
   //******************************************************************************************************
   #q_byDriveState := WORD_TO_BYTE(#ILx2T_Ref.i_woDriveStatus AND 16#000F);
   #q_xReadyToSwitchOn := #q_byDriveState = 4;
   #q_xSwitchedOn := #q_byDriveState = 6 OR #q_byDriveState = 7;
   #q_xFault := #ILx2T_Ref.stDriveStatus.FaultActive;
   #q_xWarning := #ILx2T_Ref.stDriveStatus.WarningActive;
   #q_xHALT_active := #ILx2T_Ref.stDriveStatus.HaltActive;
   #q_xRef_OK := #ILx2T_Ref.i_by_ModeStatus.%X5;
   #q_xQuickStop_Active := (#q_byDriveState = 7) AND #ILx2T_Ref.stDriveStatus.x_End;
   //******************************************************************************************************
   // MotionStat
   #q_xStandstill := #ILx2T_Ref.stDriveStatus.x_End;
   #q_xPositiveDirection := #ILx2T_Ref.i_wo_ActionWord.%X7;
   #q_xNegativeDirection := #ILx2T_Ref.i_wo_ActionWord.%X8;
   //#q_xInPositionWindow := #ILx2T_Ref.i_wo_ActionWord.%X9;
   #q_xTargetVelocityZero := #ILx2T_Ref.i_wo_ActionWord.%X11;
   #q_xAccelerating := #ILx2T_Ref.i_wo_ActionWord.%X13;
   #q_xDecelerating := #ILx2T_Ref.i_wo_ActionWord.%X12;
   #q_xConstantVelocity := #ILx2T_Ref.i_wo_ActionWord.%X14;

   #ILx2T_Ref.st_ActionWord.MotionNegative := #q_xNegativeDirection;
   //#ILx2T_Ref.st_ActionWord.InsidePosWindow := #q_xInPositionWindow;
   #ILx2T_Ref.st_ActionWord.TargetVelocityZero := #q_xTargetVelocityZero;
   #ILx2T_Ref.st_ActionWord.Decelerating := #q_xDecelerating;
   #ILx2T_Ref.st_ActionWord.Accelerating := #q_xAccelerating;
   #ILx2T_Ref.st_ActionWord.ConstantVelocity := #q_xConstantVelocity;
   #ILx2T_Ref.st_ActionWord.MotionZero := #q_xStandstill;
   #ILx2T_Ref.st_ActionWord.MotionPositive := #q_xPositiveDirection;;

   //******************************************************************************************************
   // digital Drive Inputs
   #ILx2T_Ref.x_IO_1 := #ILx2T_Ref.i_by_driveInput.%X0;
   #ILx2T_Ref.x_IO_2 := #ILx2T_Ref.i_by_driveInput.%X1;
   #ILx2T_Ref.x_IO_3 := #ILx2T_Ref.i_by_driveInput.%X2;
   #ILx2T_Ref.x_IO_4 := #ILx2T_Ref.i_by_driveInput.%X3;
   #ILx2T_Ref.x_STO_A := #ILx2T_Ref.i_by_driveInput.%X4;
   #ILx2T_Ref.x_STO_B := #ILx2T_Ref.i_by_driveInput.%X5;
   //******************************************************************************************************
   // mfStat
   #ILx2T_Ref.by_OP_ModeAct := #ILx2T_Ref.i_by_ModeStatus AND 16#0F;

   #ILx2T_Ref.st_ModeStatus.Reference_OK := #ILx2T_Ref.i_by_ModeStatus.%X5;
   #q_xRef_OK := #ILx2T_Ref.st_ModeStatus.Reference_OK;
   #ILx2T_Ref.st_ModeStatus.ModeError := #ILx2T_Ref.i_by_ModeStatus.%X6;
   #ILx2T_Ref.st_ModeStatus.ModeToggle := #ILx2T_Ref.i_by_ModeStatus.%X7;

   //******************************************************************************************************
   // Drive Control
   //******************************************************************************************************
   // Enable (Bit 8)- Disable(Bit9)
   //******************************************************************************************************
   IF #i_xDriveEnable AND #q_byDriveState > 3 AND #q_byDriveState < 9 THEN
       #ILx2T_Ref.q_wo_dmControl.%X8 := FALSE; // Disable
       #ILx2T_Ref.q_wo_dmControl.%X9 := TRUE;  // Enable
   ELSE
       #ILx2T_Ref.q_wo_dmControl.%X8 := TRUE; // Disable
       #ILx2T_Ref.q_wo_dmControl.%X9 := FALSE;  // Enable
   END_IF;
   //******************************************************************************************************
   // FAULT Reset (dmControl Bit 11)
   //******************************************************************************************************
   IF  #ILx2T_Ref.stDriveStatus.x_End AND #xQuickStopHelper THEN   // Fault Reset after QuickStop
       #ILx2T_Ref.q_wo_dmControl.%X11 := TRUE;
   ELSIF #i_xFaultReset OR #ILx2T_Ref.x_FaultResetInt THEN
       #ILx2T_Ref.q_wo_dmControl.%X11 := TRUE;
   ELSE
       #ILx2T_Ref.q_wo_dmControl.%X11 := FALSE;
   END_IF;
   //******************************************************************************************************
   // Set QuickStop
   //******************************************************************************************************
   IF #i_xQuickStop AND NOT #ILx2T_Ref.stDriveStatus.x_End THEN
       #ILx2T_Ref.q_wo_dmControl.%X10 := TRUE;
       #xQuickStopHelper := TRUE;
   ELSIF #ILx2T_Ref.x_QuickStopInt AND NOT #ILx2T_Ref.stDriveStatus.x_End THEN
       #ILx2T_Ref.q_wo_dmControl.%X10 := TRUE;
   ELSE
       #ILx2T_Ref.q_wo_dmControl.%X10 := FALSE;
   END_IF;
   // Reset QuickStopHelper
   IF #xQuickStopHelper AND #ILx2T_Ref.stDriveStatus.x_End AND #q_byDriveState <> 7 THEN
       #xQuickStopHelper := FALSE;
   END_IF;
   //******************************************************************************************************
   // Set HALT
   //******************************************************************************************************
   IF #i_xHALT THEN
       #ILx2T_Ref.q_wo_dmControl.%X13 := TRUE;
   ELSE
       #ILx2T_Ref.q_wo_dmControl.%X13 := FALSE;
       IF #q_xHALT_active THEN // Clear HALT
           #ILx2T_Ref.q_wo_dmControl.%X14 := TRUE;
       ELSE
           #ILx2T_Ref.q_wo_dmControl.%X14 := FALSE;
       END_IF;
   END_IF;
   //******************************************************************************************************
   // Continue HALT
   //******************************************************************************************************
   IF #i_xContinue THEN
       #ILx2T_Ref.q_wo_dmControl.%X15 := TRUE;
   ELSE
       #ILx2T_Ref.q_wo_dmControl.%X15 := FALSE;
   END_IF;
   //******************************************************************************************************
   // Reading Error IDs
   //******************************************************************************************************
   CASE #iState OF
       0:  // Check for error
           IF NOT #q_xFault THEN
               #q_woLastError := 0;
           END_IF;

           IF NOT #ILx2T_Ref.st_ModeStatus.ModeError THEN
               #q_woModeError := 0;
           END_IF;

           IF #q_xFault THEN
               #iState := #iState + 1;
           ELSIF #ILx2T_Ref.st_ModeStatus.ModeError THEN
               #iState := #iState + 1;
           END_IF;
           ;
       1:  // Check for parameterchannel access
           IF #ILx2T_Ref.ParChAccessID = 0 OR #ILx2T_Ref.ParChAccessID = #inAccessID THEN
               #ILx2T_Ref.ParChAccessID := #inAccessID;
               #TON_TimeOut(IN := FALSE,
                            PT := t#1s);
               #ILx2T_Ref.x_CommandReadParameter := TRUE;
               #ILx2T_Ref.udi_ModbusAddress_Read := 7178;
               #iState := #iState + 1;
           END_IF;
       2: // Start reading Last error (SopFault) 7178
           #TON_TimeOut(IN := TRUE,
                        PT := t#1s);
           IF #TON_TimeOut.Q THEN
               #TON_TimeOut(IN := FALSE,
                            PT := t#1s);
               #ILx2T_Ref.ParChAccessID := 0;
               #iErrorState := #iState;
               #iState := 100;
               // Read Done    
           ELSIF #ILx2T_Ref.x_StatusReadParameter_OK AND NOT #ILx2T_Ref.x_StatusReadParameter_Error THEN
               #TON_TimeOut(IN := FALSE,
                            PT := t#1s);
               #ILx2T_Ref.ParChAccessID := 0;
               #q_woLastError := DINT_TO_WORD(#ILx2T_Ref.di_ParameterReadValue);
               #ILx2T_Ref.x_CommandReadParameter := FALSE;
               #ILx2T_Ref.x_StatusReadParameter_OK := FALSE;
               #ILx2T_Ref.udi_ModbusAddress_Read := 0;
               #iState := #iState + 1;
               // Error response Reading
           ELSIF #ILx2T_Ref.x_StatusReadParameter_Error THEN
               #ILx2T_Ref.x_CommandReadParameter := FALSE;
               #ILx2T_Ref.x_StatusReadParameter_Error := FALSE;
               #ILx2T_Ref.udi_ModbusAddress_Read := 0;
               #TON_TimeOut(IN := FALSE,
                            PT := t#1s);
               #ILx2T_Ref.ParChAccessID := 0;
               #iErrorState := #iState;
               #iState := 100;
           END_IF;
       3:  // Check for parameterchannel access
           IF #ILx2T_Ref.ParChAccessID = 0 OR #ILx2T_Ref.ParChAccessID = #inAccessID THEN
               #ILx2T_Ref.ParChAccessID := #inAccessID;
               #TON_TimeOut(IN := FALSE,
                            PT := t#1s);
               #ILx2T_Ref.x_CommandReadParameter := TRUE;
               #ILx2T_Ref.udi_ModbusAddress_Read := 6962;
               #iState := #iState + 1;
           END_IF;
       4: // Start reading Last error (ModeError) 6962
           #TON_TimeOut(IN := TRUE,
                        PT := t#1s);
           IF #TON_TimeOut.Q THEN
               #TON_TimeOut(IN := FALSE,
                            PT := t#1s);
               #ILx2T_Ref.ParChAccessID := 0;
               #iErrorState := #iState;
               #iState := 100;
               // Read Done    
           ELSIF #ILx2T_Ref.x_StatusReadParameter_OK AND NOT #ILx2T_Ref.x_StatusReadParameter_Error THEN
               #TON_TimeOut(IN := FALSE,
                            PT := t#1s);
               #ILx2T_Ref.ParChAccessID := 0;
               #q_woModeError := DINT_TO_WORD(#ILx2T_Ref.di_ParameterReadValue);
               #ILx2T_Ref.x_CommandReadParameter := FALSE;
               #ILx2T_Ref.x_StatusReadParameter_OK := FALSE;
               #ILx2T_Ref.udi_ModbusAddress_Read := 0;
               #iState := 0;
               // Error response Reading
           ELSIF #ILx2T_Ref.x_StatusReadParameter_Error THEN
               #ILx2T_Ref.x_CommandReadParameter := FALSE;
               #ILx2T_Ref.x_StatusReadParameter_Error := FALSE;
               #ILx2T_Ref.udi_ModbusAddress_Read := 0;
               #ILx2T_Ref.ParChAccessID := 0;
               #TON_TimeOut(IN := FALSE,
                            PT := t#1s);
               #iErrorState := #iState;
               #iState := 100;
           END_IF;
       100:    // Error state        
           #iState := 0;
   END_CASE;
   //******************************************************************************************************
   // Data copy from AxisRef structure to Modbus TCP Output Data
   //******************************************************************************************************
   // Processdata
   #ILx2T_Ref.arOutputData[0] := WORD_TO_BYTE(SHR(IN := #ILx2T_Ref.q_wo_dmControl, N := 8));
   #ILx2T_Ref.arOutputData[1] := WORD_TO_BYTE(#ILx2T_Ref.q_wo_dmControl);
   #ILx2T_Ref.arOutputData[2] := WORD_TO_BYTE(SHR(IN := #ILx2T_Ref.q_dw_refA_16, N := 8));
   #ILx2T_Ref.arOutputData[3] := WORD_TO_BYTE(#ILx2T_Ref.q_dw_refA_16);
   #ILx2T_Ref.arOutputData[4] := DWORD_TO_BYTE(SHR(IN := #ILx2T_Ref.q_dw_refB_32, N := 24));
   #ILx2T_Ref.arOutputData[5] := DWORD_TO_BYTE(SHR(IN := #ILx2T_Ref.q_dw_refB_32, N := 16));
   #ILx2T_Ref.arOutputData[6] := DWORD_TO_BYTE(SHR(IN := #ILx2T_Ref.q_dw_refB_32, N := 8));
   #ILx2T_Ref.arOutputData[7] := DWORD_TO_BYTE(#ILx2T_Ref.q_dw_refB_32);
   //******************************************************************************************************
END_FUNCTION_BLOCK

FUNCTION_BLOCK "ILx2T_Homing"   // FB3, SCL
{ S7_Optimized_Access := 'TRUE' }
VERSION : 1.5
   VAR_INPUT
      i_xExecute : Bool;   // rising edge starts the operation
      i_inHM_method : Int := 33;   // Homing method (6936)
      i_diHM_p_home : DInt;   // Position at reference point after homing (10262)
      i_inHMn : Int := 60;   // Search speed - Modbus 10248
      i_inHMn_out : Int := 6;   // move out speed - Modbus 10250
      i_diHMdisusr : DInt := 200;   // Distance from switching edge to reference point - Modbus 10254
      i_diHMoutdisusr : DInt;   // Max. distance for search for switching edge - Modbus 10252
      i_diHMsrchdisusr : DInt;   // Max. search distance after overrun of switch - Modbus 10266
   END_VAR
   VAR_OUTPUT
      q_xDone : Bool;   // reference movement finished without error
      q_xError : Bool;   // finished with error
      q_xCommandAborted : Bool;   // function aborted
      q_xBusy : Bool;   // function is active
   END_VAR
   VAR_IN_OUT
      ILx2T_Ref : "ILx2T_Ref";   // Axis reference structure
   END_VAR
   VAR
      inState : Int;   // internal state machine
      inAccessID : Int;   // own access ID
      inErrorState : Int;
      woInternalErrorID : Word;   // internal FB error ID
      xModeToggleHelper : Bool;
      TON_Timeout : TON_TIME;
      inHelperState : Int;
      diHelperParameterValue : DInt;
      udiHelperParameterAddress : UDInt;
   END_VAR
BEGIN
   // *******************************************************************************
   // Init after Restart
   // *******************************************************************************
   // Check for PLC restart (1st call of this FB)
   IF #inAccessID = 0 THEN
       #ILx2T_Ref.InitAccessID := #ILx2T_Ref.InitAccessID + 1;
       #inAccessID := #ILx2T_Ref.InitAccessID;
   END_IF;

   CASE #inState OF
           // ******************************************************************************************************
       0:  // idle state
           IF #i_xExecute THEN
               #q_xBusy := TRUE;
               #inErrorState := 0;
               #woInternalErrorID := 0;
               #inState := #inState + 1;
           ELSE
               #q_xDone := FALSE;
               #q_xError := FALSE;
               #q_xBusy := FALSE;
               #q_xCommandAborted := FALSE;
           END_IF;
           // ******************************************************************************************************
       1:  // Check for drive state and access ID
           IF NOT #ILx2T_Ref.stDriveStatus.x_End AND #ILx2T_Ref.by_OP_ModeAct <> 2 THEN  // A318 operating mode active
               #q_xError := TRUE;
               #woInternalErrorID := 16#A318;
               #inErrorState := #inState;
               #inState := 100;
           ELSIF ((#ILx2T_Ref.i_woDriveStatus AND 16#F) = 6) OR ((#ILx2T_Ref.i_woDriveStatus AND 16#F) = 7) THEN
               IF #i_inHM_method = 35 THEN
                   #inState := 8;
               ELSE
                   #inState := #inState + 1;
               END_IF;
           ELSE
               #q_xError := TRUE;
               #inErrorState := #inState;
               #inState := 100;
           END_IF;
           // ******************************************************************************************************
       2:  // Wtrite Parameter 10262 (32 Bit) - homing position
           #udiHelperParameterAddress := 10262;
           #diHelperParameterValue := #i_diHM_p_home;
           #inHelperState := #inState + 1;
           #inState := 50;
           // ******************************************************************************************************
       3:  // Wtrite Parameter 10248 (16 Bit) - HMn search speed
           #udiHelperParameterAddress := 10248;
           #diHelperParameterValue := #i_inHMn;
           #inHelperState := #inState + 1;
           #inState := 50;
           // ******************************************************************************************************
       4:  // Wtrite Parameter 10250 (16 Bit) - HMn_out move out speed
           #udiHelperParameterAddress := 10250;
           #diHelperParameterValue := #i_inHMn_out;
           #inHelperState := #inState + 1;
           #inState := 50;
           // ******************************************************************************************************
       5:  // Wtrite Parameter 10254 (32 Bit) - HM_disusr - distance from switching edge
           #udiHelperParameterAddress := 10254;
           #diHelperParameterValue := #i_diHMdisusr;
           #inHelperState := #inState + 1;
           #inState := 50;
           // ******************************************************************************************************
       6:  // Wtrite Parameter 10252 (32 Bit) - HM_outdisusr - max. search distance from switching edge
           #udiHelperParameterAddress := 10252;
           #diHelperParameterValue := #i_diHMoutdisusr;
           #inHelperState := #inState + 1;
           #inState := 50;
           // ******************************************************************************************************
       7:  // Wtrite Parameter 10266 (32 Bit) - HM_srchdisusr - max. search distance 
           #udiHelperParameterAddress := 10266;
           #diHelperParameterValue := #i_diHMsrchdisusr;
           #inHelperState := #inState + 1;
           #inState := 50;
           // ******************************************************************************************************
           // Start Homing
           // ******************************************************************************************************
       8: // Start Homing via Processchannel
           //   Mode 02 hex = Dimension Setting (RefA16 = not used / RefB32 = reference position)
           //   Mode 12 hex = Reference movement (RefA16 = homing mode / RefB32 = not used)
           CASE #i_inHM_method OF
               35: // type SetPosition
                   #ILx2T_Ref.q_wo_dmControl := #ILx2T_Ref.q_wo_dmControl AND 16#FF80;
                   #ILx2T_Ref.q_wo_dmControl := #ILx2T_Ref.q_wo_dmControl OR 16#0002;
                   #ILx2T_Ref.q_dw_refA_16 := 0;
                   #ILx2T_Ref.q_dw_refB_32 := DINT_TO_WORD(#i_diHM_p_home);
                   #inState := #inState + 1;
               0..34:
                   #ILx2T_Ref.q_wo_dmControl := #ILx2T_Ref.q_wo_dmControl AND 16#FF80;
                   #ILx2T_Ref.q_wo_dmControl := #ILx2T_Ref.q_wo_dmControl OR 16#0012;
                   #ILx2T_Ref.q_dw_refA_16 := INT_TO_WORD(#i_inHM_method);
                   #ILx2T_Ref.q_dw_refB_32 := 0;
                   #inState := #inState + 1;
               ELSE
                   #inErrorState := #inState;
                   #inState := 100;
           END_CASE;
           // ******************************************************************************************************
       9: // Mode Toggle
           #xModeToggleHelper := NOT #ILx2T_Ref.st_ModeStatus.ModeToggle;  // save toggle bit 
           IF #ILx2T_Ref.st_ModeStatus.ModeToggle THEN
               #ILx2T_Ref.q_wo_dmControl := #ILx2T_Ref.q_wo_dmControl AND 16#FF7F;
           ELSE
               #ILx2T_Ref.q_wo_dmControl := #ILx2T_Ref.q_wo_dmControl OR 16#0080;
           END_IF;
           #inState := #inState + 1;
           // ******************************************************************************************************
       10: // Check for mode toggle and number of operating mode OK
           IF NOT (#xModeToggleHelper XOR #ILx2T_Ref.st_ModeStatus.ModeToggle) AND (#ILx2T_Ref.by_OP_ModeAct = 16#0002) THEN                            // Check operating mode number
               #TON_Timeout(IN := FALSE,
                            PT := t#1s);
               #inState := #inState + 1;  // Command OK
           ELSE
               // TIMEOUT ERROR
               #TON_Timeout(IN := TRUE,
                            PT := t#1s);
               IF #TON_Timeout.Q THEN
                   #TON_Timeout(IN := FALSE,
                                PT := t#1s);
                   #q_xError := TRUE;
                   #inErrorState := #inState;
                   #inState := 100;
               END_IF;
           END_IF;
           // ******************************************************************************************************
       11: // Check operating mode
           // Mode OK -> Check drive status (x_Add, x_End and x_Error)
           IF #ILx2T_Ref.st_ModeStatus.Reference_OK AND #ILx2T_Ref.stDriveStatus.x_End AND NOT #ILx2T_Ref.stDriveStatus.x_Err THEN  // finished without Error     
               #q_xBusy := FALSE;
               #q_xDone := TRUE;
               #inState := 110;
               //ELSIF NOT #ILx2T_Ref.stDriveStatus.x_End AND NOT #ILx2T_Ref.stDriveStatus.x_Err THEN  // Mode sill active     
               //    ;
           ELSIF #ILx2T_Ref.stDriveStatus.x_End AND #ILx2T_Ref.stDriveStatus.x_Err THEN  // finished with Error     
               #inErrorState := #inState;
               #inState := 100;
           ELSIF #ILx2T_Ref.by_OP_ModeAct <> 16#0002 THEN   // check for correct operating mode number
               #q_xCommandAborted := TRUE;
               #q_xBusy := FALSE;
               #q_xDone := FALSE;
               #inState := 110;
           END_IF;
           // ******************************************************************************************************
           // Parameter channel handling
           // ******************************************************************************************************
       50: // Check for parameterchannel access
           IF #ILx2T_Ref.ParChAccessID = 0 OR #ILx2T_Ref.ParChAccessID = #inAccessID THEN
               #ILx2T_Ref.ParChAccessID := #inAccessID;   // grab access to parameter channel
               #TON_Timeout(IN := FALSE,
                            PT := t#1s);
               #ILx2T_Ref.x_CommandWriteParameter := TRUE;
               #ILx2T_Ref.udi_ModbusAddress_Write := #udiHelperParameterAddress;
               #ILx2T_Ref.di_ParameterWriteValue := #diHelperParameterValue;
               #inState := #inState + 1;
           END_IF;
       51: // Check for Parameterchannel response
           #TON_Timeout(IN := TRUE,
                        PT := t#1s);
           IF #TON_Timeout.Q THEN
               #TON_Timeout(IN := FALSE,
                            PT := t#1s);
               #q_xError := TRUE;
               #ILx2T_Ref.ParChAccessID := 0;   // release access to parameter channel
               #inErrorState := #inState;
               #inState := 100;
               // Write Done    
           ELSIF #ILx2T_Ref.x_Status_WriteParameter_OK AND NOT #ILx2T_Ref.x_Status_WriteParameter_Error THEN
               #TON_Timeout(IN := FALSE,
                            PT := t#1s);
               #ILx2T_Ref.di_ParameterWriteValue := 0;
               #ILx2T_Ref.x_CommandWriteParameter := FALSE;
               #ILx2T_Ref.x_Status_WriteParameter_OK := FALSE;
               #ILx2T_Ref.udi_ModbusAddress_Write := 0;
               #ILx2T_Ref.ParChAccessID := 0;   // release access to parameter channel
               #inState := #inHelperState;
               // Error response Writing
           ELSIF #ILx2T_Ref.x_Status_WriteParameter_Error THEN
               #ILx2T_Ref.x_CommandWriteParameter := FALSE;
               #ILx2T_Ref.x_Status_WriteParameter_Error := FALSE;
               #ILx2T_Ref.udi_ModbusAddress_Write := 0;
               #TON_Timeout(IN := FALSE,
                            PT := t#1s);
               #ILx2T_Ref.ParChAccessID := 0;   // release access to parameter channel
               #inErrorState := #inState;
               #inState := 100;
           END_IF;
           // ******************************************************************************************************
       100:  // Error state
           IF #ILx2T_Ref.ParChAccessID = #inAccessID THEN
               #ILx2T_Ref.ParChAccessID := 0;   // grab access to parameter channel
           END_IF;
           IF #ILx2T_Ref.ProChAccessID = #inAccessID THEN
               #ILx2T_Ref.ProChAccessID := 0;   // grab access to parameter channel
           END_IF;
           #q_xBusy := FALSE;
           #q_xError := TRUE;
           #inState := 110;
           // ******************************************************************************************************
       110:  // finished
           IF NOT #i_xExecute THEN
               #q_xDone := FALSE;
               #q_xError := FALSE;
               #q_xBusy := FALSE;
               #q_xCommandAborted := FALSE;
               #inState := 0;
           END_IF;
           // ******************************************************************************************************
   END_CASE;
END_FUNCTION_BLOCK

FUNCTION_BLOCK "ILx2T_Jog"   // FB4, SCL
{ S7_Optimized_Access := 'TRUE' }
VERSION : 1.5
   VAR_INPUT
      i_xForward : Bool;   // Jog forward
      i_xBackward : Bool;   // Jog backward
      i_xFast : Bool;   // Jog fast
   END_VAR
   VAR_OUTPUT
      q_xError : Bool;   // finished with error
      q_xCommandAborted : Bool;   // function aborted
      q_xBusy : Bool;   // function is busy
   END_VAR
   VAR_IN_OUT
      ILx2T_Ref : "ILx2T_Ref";   // Axis reference structure
   END_VAR
   VAR
      inState : Int;   // internal state machine
      inAccessID : Int;   // own access ID
      inHelperState : Int;
      inErrorState : Int;
      woInternalErrorID : Word;   // internal FB error ID
      xModeToggleHelper : Bool;
      xHelperForward : Bool;
      xHelperBackward : Bool;
      xHelperFast : Bool;
      TON_Timeout : TON_TIME;
   END_VAR
BEGIN
   // *******************************************************************************
   // Init after Restart
   // *******************************************************************************
   // Check for PLC restart (1st call of this FB)
   IF #inAccessID = 0 THEN
       #ILx2T_Ref.InitAccessID := #ILx2T_Ref.InitAccessID + 1;
       #inAccessID := #ILx2T_Ref.InitAccessID;
   END_IF;

   CASE #inState OF
           // ******************************************************************************************************
       0:  // idle state
           IF #i_xForward XOR #i_xBackward THEN
               #xHelperForward := #i_xForward;
               #xHelperBackward := #i_xBackward;
               #xHelperFast := #i_xFast;
               #q_xBusy := TRUE;
               #inErrorState := 0;
               #inState := #inState + 1;
           ELSE
               #q_xError := FALSE;
               #q_xBusy := FALSE;
               #q_xCommandAborted := FALSE;
           END_IF;
           // ******************************************************************************************************
       1:  // Check for drive state and access ID
           IF NOT #ILx2T_Ref.stDriveStatus.x_End AND #ILx2T_Ref.by_OP_ModeAct <> 1 THEN  // A318 operating mode active
               #q_xError := TRUE;
               #woInternalErrorID := 16#A318;
               #inErrorState := #inState;
               #inState := 100;
           ELSIF ((#ILx2T_Ref.i_woDriveStatus AND 16#0F) = 16#06) OR ((#ILx2T_Ref.i_woDriveStatus AND 16#0F) = 16#07) THEN
               IF #ILx2T_Ref.ProChAccessID = 0 OR #ILx2T_Ref.ProChAccessID = #inAccessID THEN
                   #ILx2T_Ref.ProChAccessID := #inAccessID;   // grab access to proccessdata channel
                   // Start Movement via Processchannel
                   // Mode 01 hex = Jog mode (RefA16 = jog activate / RefB32 = reserved)
                   #ILx2T_Ref.q_dw_refB_32 := 0;
                   IF NOT #xHelperForward AND NOT #xHelperBackward THEN
                       #ILx2T_Ref.q_dw_refA_16 := 16#00;
                   ELSIF #xHelperForward AND NOT #xHelperFast THEN
                       #ILx2T_Ref.q_dw_refA_16 := 16#01;
                   ELSIF #xHelperBackward AND NOT #xHelperFast THEN
                       #ILx2T_Ref.q_dw_refA_16 := 16#02;
                   ELSIF #xHelperForward AND #xHelperFast THEN
                       #ILx2T_Ref.q_dw_refA_16 := 16#05;
                   ELSIF #xHelperBackward AND #xHelperFast THEN
                       #ILx2T_Ref.q_dw_refA_16 := 16#06;
                   END_IF;
                   #ILx2T_Ref.q_wo_dmControl := #ILx2T_Ref.q_wo_dmControl AND 16#FF80;
                   #ILx2T_Ref.q_wo_dmControl := #ILx2T_Ref.q_wo_dmControl OR 16#0001;
                   #inState := #inState + 1;
               END_IF;
           ELSE
               #q_xError := TRUE;
               #inErrorState := #inState;
               #inState := 100;
           END_IF;
           // ******************************************************************************************************
       2: // Mode Toggle
           #xModeToggleHelper := NOT #ILx2T_Ref.st_ModeStatus.ModeToggle;  // save toggle bit 
           IF NOT #xModeToggleHelper THEN
               #ILx2T_Ref.q_wo_dmControl := #ILx2T_Ref.q_wo_dmControl AND 16#FF7F;
           ELSE
               #ILx2T_Ref.q_wo_dmControl := #ILx2T_Ref.q_wo_dmControl OR 16#0080;
           END_IF;
           #inState := #inState + 1;
           // ******************************************************************************************************
       3: // Check for mode response OK
           // Check for mode toggle and number of operating mode OK
           IF NOT (#xModeToggleHelper XOR #ILx2T_Ref.st_ModeStatus.ModeToggle) AND (#ILx2T_Ref.by_OP_ModeAct = 16#01) THEN                            // Check operating mode number
               #TON_Timeout(IN := FALSE,
                            PT := t#1s);
               #ILx2T_Ref.ProChAccessID := 0;   // release access to proccessdata channel
               #inState := #inState + 1;
           ELSE
               // TIMEOUT ERROR
               #TON_Timeout(IN := TRUE,
                            PT := t#1s);
               IF #TON_Timeout.Q THEN
                   #TON_Timeout(IN := FALSE,
                                PT := t#1s);
                   #q_xError := TRUE;
                   #inErrorState := #inState;
                   #inState := 100;
               END_IF;
           END_IF;
           // ******************************************************************************************************
       4: // Check operating mode
           // x_Error
           IF #ILx2T_Ref.stDriveStatus.x_Err THEN  // error     
               #inErrorState := #inState;
               #inState := 100;
               // Monitoring of actual operating mode
           ELSIF (#ILx2T_Ref.by_OP_ModeAct <> 16#01) THEN
               #q_xCommandAborted := TRUE;
               #q_xBusy := FALSE;
               #inState := 110;
               // Check if command has changed
               // x_END and no command 
           ELSIF #ILx2T_Ref.stDriveStatus.x_End AND NOT #xHelperForward AND NOT #xHelperBackward THEN  // error     
               #q_xBusy := FALSE;
               #inState := 0;
           ELSIF NOT (#i_xBackward XOR #i_xForward) THEN
               #xHelperForward := FALSE;
               #xHelperBackward := FALSE;
               #xHelperFast := FALSE;
               #inState := 1;
           ELSIF #xHelperForward <> #i_xForward THEN
               #inState := 0;
           ELSIF #xHelperBackward <> #i_xBackward THEN
               #inState := 0;
           ELSIF #xHelperFast <> #i_xFast THEN
               #inState := 0;
           END_IF;

           // ******************************************************************************************************
       100:  // Error state
           IF #ILx2T_Ref.ProChAccessID = #inAccessID THEN
               #ILx2T_Ref.ProChAccessID := 0;   // release access to proccessdata channel
           END_IF;
           #q_xBusy := FALSE;
           #q_xError := TRUE;
           #inState := 110;
           // ******************************************************************************************************
       110:  // finished
           IF NOT #i_xForward AND NOT #i_xBackward THEN
               #q_xError := FALSE;
               #q_xBusy := FALSE;
               #q_xCommandAborted := FALSE;
               #inState := 0;
           END_IF;
           // ******************************************************************************************************
   END_CASE;
END_FUNCTION_BLOCK

FUNCTION_BLOCK "ILx2T_Parameter_Read_Write"   // FB5, SCL
{ S7_Optimized_Access := 'TRUE' }
VERSION : 1.5
   VAR_INPUT
      i_xParameterRead : Bool;   // TRUE = Reading value continuously
      i_xParameterWrite : Bool;   // rising edge = Writing once
      i_woParameterAddress : Word;   // Parameter address (see product manual)
      i_byWriteParameterLength : Byte;   // parameter length in bytes ( 2 or 4 bytes)
      i_diWriteParameterValue : DInt;   // parameter write value
   END_VAR
   VAR_OUTPUT
      q_xReadValueValid : Bool;   // reading value is valid
      q_xWriteDone : Bool;   // writing finished without error
      q_xError : Bool;   // finished with error
      q_xBusy : Bool;   // function is active
      q_diReadParameterValue : DInt;   // reading value
   END_VAR
   VAR_IN_OUT
      ILx2T_Ref : "ILx2T_Ref";   // Axis reference structure
   END_VAR
   VAR
      inState : Int;   // internal state machine
      inAccessID : Int;   // own access ID
      inErrorState : Int;
      dwParaChErrorNo : DWord;   // parameter channe error ID
      xHelperWrite : Bool;
      xHelperRead : Bool;
      TON_Timeout : TON_TIME;
   END_VAR
BEGIN
   // *******************************************************************************
   // Init after Restart
   // *******************************************************************************
   // Check for PLC restart (1st call of this FB)
   IF #inAccessID = 0 THEN
       #ILx2T_Ref.InitAccessID := #ILx2T_Ref.InitAccessID + 1;
       #inAccessID := #ILx2T_Ref.InitAccessID;
   END_IF;

   CASE #inState OF
           // ******************************************************************************************************
       0:  // idle state
           IF #i_xParameterWrite XOR #i_xParameterRead THEN
               #xHelperWrite := #i_xParameterWrite;
               #xHelperRead := #i_xParameterRead;
               #q_xBusy := TRUE;
               #inErrorState := 0;
               #dwParaChErrorNo := 0;
               #inState := #inState + 1;
           ELSE
               #q_xWriteDone := FALSE;
               #q_xError := FALSE;
               #q_xBusy := FALSE;
               #q_xReadValueValid := FALSE;
               #q_diReadParameterValue := 0;
           END_IF;
           // ******************************************************************************************************
       1:  // Check for parameterchannel access
           IF #ILx2T_Ref.ParChAccessID = 0 OR #ILx2T_Ref.ParChAccessID = #inAccessID THEN
               #ILx2T_Ref.ParChAccessID := #inAccessID;   // grab access to parameter channel
               #inState := #inState + 1;
           END_IF;
           // ******************************************************************************************************
       2:// Prepare parameterchannel command
           #TON_Timeout(IN := FALSE,
                        PT := t#1s);
           IF #xHelperRead THEN
               #ILx2T_Ref.x_CommandReadParameter := TRUE;
               #ILx2T_Ref.udi_ModbusAddress_Read := #i_woParameterAddress;
               #inState := #inState + 1;
           ELSIF #xHelperWrite THEN
               #ILx2T_Ref.x_CommandWriteParameter := TRUE;
               #ILx2T_Ref.udi_ModbusAddress_Write := #i_woParameterAddress;
               #ILx2T_Ref.di_ParameterWriteValue := #i_diWriteParameterValue;
               #inState := #inState + 1;
           END_IF;
           // ******************************************************************************************************
       3: // Check for Parameterchannel response
           #TON_Timeout(IN := TRUE,
                        PT := t#1s);
           IF #TON_Timeout.Q THEN
               #TON_Timeout(IN := FALSE,
                            PT := t#1s);
               #q_xError := TRUE;
               #inErrorState := #inState;
               #inState := 100;
               // Read Done    
           ELSIF #xHelperRead AND #ILx2T_Ref.x_StatusReadParameter_OK AND NOT #ILx2T_Ref.x_StatusReadParameter_Error THEN
               #TON_Timeout(IN := FALSE,
                            PT := t#1s);
               #q_diReadParameterValue := #ILx2T_Ref.di_ParameterReadValue;
               #q_xReadValueValid := TRUE;
               #ILx2T_Ref.x_CommandReadParameter := FALSE;
               #ILx2T_Ref.x_StatusReadParameter_OK := FALSE;
               #ILx2T_Ref.udi_ModbusAddress_Read := 0;
               #inState := #inState + 1;
               // Write Done    
           ELSIF #xHelperWrite AND #ILx2T_Ref.x_Status_WriteParameter_OK AND NOT #ILx2T_Ref.x_Status_WriteParameter_Error THEN
               #TON_Timeout(IN := FALSE,
                            PT := t#1s);
               #ILx2T_Ref.di_ParameterWriteValue := 0;
               #q_xWriteDone := TRUE;
               #ILx2T_Ref.x_CommandWriteParameter := FALSE;
               #ILx2T_Ref.x_Status_WriteParameter_OK := FALSE;
               #ILx2T_Ref.udi_ModbusAddress_Write := 0;
               #inState := #inState + 1;
               // Error response Reading
           ELSIF #ILx2T_Ref.x_StatusReadParameter_Error THEN
               #ILx2T_Ref.x_CommandReadParameter := FALSE;
               #ILx2T_Ref.x_StatusReadParameter_Error := FALSE;
               #ILx2T_Ref.udi_ModbusAddress_Read := 0;
               #TON_Timeout(IN := FALSE,
                            PT := t#1s);
               #inErrorState := #inState;
               #inState := 100;
               // Error response Writing
           ELSIF #ILx2T_Ref.x_Status_WriteParameter_Error THEN
               #ILx2T_Ref.x_CommandWriteParameter := FALSE;
               #ILx2T_Ref.x_Status_WriteParameter_Error := FALSE;
               #ILx2T_Ref.udi_ModbusAddress_Write := 0;
               #TON_Timeout(IN := FALSE,
                            PT := t#1s);
               #inErrorState := #inState;
               #inState := 100;
           END_IF;
           // ******************************************************************************************************
       4:  // Check for Parameterchannel in idle state
           #TON_Timeout(IN := TRUE,
                        PT := t#1s);
           IF #TON_Timeout.Q THEN
               #TON_Timeout(IN := FALSE,
                            PT := t#1s);
               #q_xError := TRUE;
               #inErrorState := #inState;
               #inState := 100;
           ELSIF NOT #ILx2T_Ref.x_StatusReadParameter_OK AND NOT #ILx2T_Ref.x_StatusReadParameter_Error
               AND NOT #ILx2T_Ref.x_Status_WriteParameter_OK AND NOT #ILx2T_Ref.x_Status_WriteParameter_Error THEN
               #ILx2T_Ref.ParChAccessID := 0;   // grab access to parameter channel
               #TON_Timeout(IN := FALSE,
                            PT := t#1s);
               IF #xHelperWrite THEN
                   #q_xBusy := FALSE;
                   #inState := 110;
               ELSE
                   #inState := 0;
               END_IF;
           END_IF;
       100:  // Error state
           IF #ILx2T_Ref.ParChAccessID = #inAccessID THEN
               #ILx2T_Ref.ParChAccessID := 0;   // release access to proccessdata channel
           END_IF;
           #q_xBusy := FALSE;
           #q_xError := TRUE;
           #inState := 110;
           // ******************************************************************************************************
       110:  // finished
           IF NOT #i_xParameterWrite AND NOT #i_xParameterRead THEN
               #q_xWriteDone := FALSE;
               #q_xError := FALSE;
               #q_xBusy := FALSE;
               #q_xReadValueValid := FALSE;
               #q_diReadParameterValue := 0;
               #inState := 0;
           END_IF;
           // ******************************************************************************************************
   END_CASE;
END_FUNCTION_BLOCK

FUNCTION_BLOCK "ILx2T_ProfilePosition"   // FB6, SCL
{ S7_Optimized_Access := 'TRUE' }
VERSION : 1.5
   VAR_INPUT
      i_xExecute : Bool;   // rising edge starts a new movement
      i_xAbort : Bool;   // abort active movement
      i_inPTP_Type : Int;   // 1=absolute / 2=additive / 3=relative
      i_diTargetPosition : DInt;   // Target position value
      i_inTargetVelocity : Int;   // Target velocity value
   END_VAR
   VAR_OUTPUT
      q_xDone : Bool;   // Target position reached
      q_xError : Bool;   // finished with error
      q_xCommandAborted : Bool;   // function aborted
      q_xBusy : Bool;   // function is active
   END_VAR
   VAR_IN_OUT
      ILx2T_Ref : "ILx2T_Ref";   // Axis reference structure
   END_VAR
   VAR
      inState : Int;   // internal state machine
      inAccessID : Int;   // own access ID
      inHelperState : Int;
      inErrorState : Int;
      woInternalErrorID : Word;   // internal FB error ID
      xModeToggleHelper : Bool;
      xHelperExecute : Bool;
      inHelperTargetVelocity : Int;
      TON_Timeout : TON_TIME;
   END_VAR
BEGIN
   // *******************************************************************************
   // Init after Restart
   // *******************************************************************************
   // Check for PLC restart (1st call of this FB)
   IF #inAccessID = 0 THEN
       #ILx2T_Ref.InitAccessID := #ILx2T_Ref.InitAccessID + 1;
       #inAccessID := #ILx2T_Ref.InitAccessID;
   END_IF;

   CASE #inState OF
           // ******************************************************************************************************
       0:  // idle state
           IF #i_xExecute THEN
               #q_xBusy := TRUE;
               #inErrorState := 0;
               #inState := #inState + 1;
           ELSE
               #q_xDone := FALSE;
               #q_xError := FALSE;
               #q_xBusy := FALSE;
               #q_xCommandAborted := FALSE;
           END_IF;
           // ******************************************************************************************************
       1:  // Check for drive state and access ID
           IF NOT #ILx2T_Ref.stDriveStatus.x_End AND #ILx2T_Ref.by_OP_ModeAct <> 3 THEN  // A318 operating mode active
               #q_xError := TRUE;
               #woInternalErrorID := 16#A318;
               #inErrorState := #inState;
               #inState := 100;
           ELSIF (#ILx2T_Ref.i_woDriveStatus AND 16#F) = 6 THEN
               #inState := #inState + 1;
           ELSE
               #q_xError := TRUE;
               #inErrorState := #inState;
               #inState := 100;
           END_IF;
           // ******************************************************************************************************
       2: // Start Movement via Processchannel
           //   i_inPTP_Type 1 = Mode 03 hex = move absolute (RefA32 = target velocity / RefB32 = target position)
           //   i_inPTP_Type 2 = Mode 13 hex = move additive (RefA32 = target velocity / RefB32 = target position)
           //   i_inPTP_Type 3 = Mode 23 hex = move relative (RefA32 = target velocity / RefB32 = target position)
           #ILx2T_Ref.q_dw_refA_16 := INT_TO_WORD(#i_inTargetVelocity);
           #inHelperTargetVelocity := #i_inTargetVelocity;
           #ILx2T_Ref.q_dw_refB_32 := DINT_TO_DWORD(#i_diTargetPosition);
           #xHelperExecute := FALSE;
           CASE #i_inPTP_Type OF
               1: // Move absolute
                   #ILx2T_Ref.q_wo_dmControl := #ILx2T_Ref.q_wo_dmControl AND 16#FF80;
                   #ILx2T_Ref.q_wo_dmControl := #ILx2T_Ref.q_wo_dmControl OR 16#0003;
                   #inState := #inState + 1;
               2: // Move additive
                   #ILx2T_Ref.q_wo_dmControl := #ILx2T_Ref.q_wo_dmControl AND 16#FF80;
                   #ILx2T_Ref.q_wo_dmControl := #ILx2T_Ref.q_wo_dmControl OR 16#0013;
                   #inState := #inState + 1;
               3: // Move relative
                   #ILx2T_Ref.q_wo_dmControl := #ILx2T_Ref.q_wo_dmControl AND 16#FF80;
                   #ILx2T_Ref.q_wo_dmControl := #ILx2T_Ref.q_wo_dmControl OR 16#0023;
                   #inState := #inState + 1;
               ELSE
                   #inErrorState := #inState;
                   #inState := 100;
           END_CASE;

           // ******************************************************************************************************
       3: // ModeToggle 
           IF NOT #i_xExecute THEN
               #xHelperExecute := TRUE;
           END_IF;
           #xModeToggleHelper := NOT #ILx2T_Ref.st_ModeStatus.ModeToggle;  // save toggle bit 
           IF NOT #xModeToggleHelper THEN
               #ILx2T_Ref.q_wo_dmControl := #ILx2T_Ref.q_wo_dmControl AND 16#FF7F;
           ELSE
               #ILx2T_Ref.q_wo_dmControl := #ILx2T_Ref.q_wo_dmControl OR 16#0080;
           END_IF;
           #inState := #inState + 1;
           // ******************************************************************************************************
       4: // Check for mode toggle and number of operating mode OK
           IF NOT #i_xExecute THEN
               #xHelperExecute := TRUE;
           END_IF;
           IF NOT (#xModeToggleHelper XOR #ILx2T_Ref.st_ModeStatus.ModeToggle) AND (#ILx2T_Ref.by_OP_ModeAct = 16#0003) THEN                            // Check operating mode number
               #TON_Timeout(IN := FALSE,
                            PT := t#1s);
               #inState := #inState + 1;  // Command OK
           ELSE
               // TIMEOUT ERROR
               #TON_Timeout(IN := TRUE,
                            PT := t#1s);
               IF #TON_Timeout.Q THEN
                   #TON_Timeout(IN := FALSE,
                                PT := t#1s);
                   #q_xError := TRUE;
                   #inErrorState := #inState;
                   #inState := 100;
               END_IF;
           END_IF;
           // ******************************************************************************************************
       5: // Check operating mode
           IF NOT #i_xExecute THEN
               #xHelperExecute := TRUE;
           END_IF;
           // Mode OK -> Check drive status (x_Add, x_End and x_Error)
           IF #ILx2T_Ref.stDriveStatus.x_Add AND #ILx2T_Ref.stDriveStatus.x_End AND NOT #ILx2T_Ref.stDriveStatus.x_Err THEN  // finished without Error     
               #q_xBusy := FALSE;
               #q_xDone := TRUE;
               #inState := 110;
           ELSIF #ILx2T_Ref.stDriveStatus.x_End AND #ILx2T_Ref.stDriveStatus.x_Err THEN  // finished with Error     
               #inErrorState := #inState;
               #inState := 100;
           ELSIF #ILx2T_Ref.by_OP_ModeAct <> 16#0003 THEN   // check for correct operating mode number
               #q_xCommandAborted := TRUE;
               #q_xBusy := FALSE;
               #q_xDone := FALSE;
               #inState := 110;
           ELSIF #i_xExecute AND #xHelperExecute THEN
               #inState := 2;
           ELSIF #i_xAbort THEN
               #ILx2T_Ref.x_QuickStopInt := TRUE;
               #inState := #inState + 1;
           // Velocity can be changed during movement (only move absolute)
           ELSIF #i_inPTP_Type = 1 THEN
               IF #inHelperTargetVelocity <> #i_inTargetVelocity THEN
                   #inState := 2;
               END_IF;
           END_IF;
       6:
           IF #ILx2T_Ref.stDriveStatus.x_End AND (#ILx2T_Ref.i_woDriveStatus AND 16#F) >= 7 THEN  // Check for STANDSTILL
               #ILx2T_Ref.x_QuickStopInt := FALSE;
               #ILx2T_Ref.x_FaultResetInt := TRUE;
               #TON_Timeout(IN := TRUE,
                            PT := t#1s);
               IF #TON_Timeout.Q THEN
                   #TON_Timeout(IN := FALSE,
                                PT := t#1s);
                   #ILx2T_Ref.x_FaultResetInt := FALSE;
                   #q_xError := TRUE;
                   #inErrorState := #inState;
                   #inState := 100;
               END_IF;
           ELSIF #ILx2T_Ref.stDriveStatus.x_End AND (#ILx2T_Ref.i_woDriveStatus AND 16#F) < 7 THEN  // Check for STANDSTILL
               #ILx2T_Ref.x_QuickStopInt := FALSE;
               #ILx2T_Ref.x_FaultResetInt := FALSE;
               #q_xCommandAborted := TRUE;
               #q_xBusy := FALSE;
               #q_xDone := FALSE;
               #inState := 110;
           END_IF;

           // ******************************************************************************************************
       100:  // Error state
           #q_xBusy := FALSE;
           #q_xError := TRUE;
           #inState := 110;
           // ******************************************************************************************************
       110:  // finished
           IF NOT #i_xExecute AND NOT #i_xAbort THEN
               #q_xDone := FALSE;
               #q_xError := FALSE;
               #q_xBusy := FALSE;
               #q_xCommandAborted := FALSE;
               #inState := 0;
           END_IF;
           // ******************************************************************************************************
   END_CASE;
END_FUNCTION_BLOCK

FUNCTION_BLOCK "ILx2T_ProfileVelocity"   // FB8, SCL
{ S7_Optimized_Access := 'TRUE' }
VERSION : 1.5
   VAR_INPUT
      i_xExecute : Bool;   // Start movement
      i_xAbort : Bool;   // Abort current movement
      i_inTargetVelocity : Int;   // Target speed
   END_VAR
   VAR_OUTPUT
      q_xTargetVelocityReached : Bool;   // Target velocity reached
      q_xError : Bool;   // FB finished with error
      q_xCommandAborted : Bool;   // FB aborted
      q_xBusy : Bool;   // function block is busy
   END_VAR
   VAR_IN_OUT
      ILx2T_Ref : "ILx2T_Ref";   // Axis reference structure
   END_VAR
   VAR
      inState : Int;   // internal state machine
      inAccessID : Int;   // own access ID
      inHelperState : Int;
      inErrorState : Int;
      woInternalErrorID : Word;   // internal FB error ID
      xModeToggleHelper : Bool;
      inTargetVelocityHelper : Int;
      TON_Timeout : TON_TIME;
   END_VAR
BEGIN
   // *******************************************************************************
   // Init after Restart
   // *******************************************************************************
   // Check for PLC restart (1st call of this FB)
   IF #inAccessID = 0 THEN
       #ILx2T_Ref.InitAccessID := #ILx2T_Ref.InitAccessID + 1;
       #inAccessID := #ILx2T_Ref.InitAccessID;
   END_IF;

   CASE #inState OF
           // ******************************************************************************************************
       0:  // idle state
           IF #i_xExecute THEN
               #q_xBusy := TRUE;
               #inErrorState := 0;
               #inState := #inState + 1;
           ELSE
               #q_xTargetVelocityReached := FALSE;
               #q_xError := FALSE;
               #q_xBusy := FALSE;
               #q_xCommandAborted := FALSE;
           END_IF;
           // ******************************************************************************************************
       1:  // Check for drive state and access ID
           IF NOT #ILx2T_Ref.stDriveStatus.x_End AND #ILx2T_Ref.by_OP_ModeAct <> 4 THEN  // A318 operating mode active
               #q_xError := TRUE;
               #woInternalErrorID := 16#A318;
               #inErrorState := #inState;
               #inState := 100;
           ELSIF (#ILx2T_Ref.i_woDriveStatus AND 16#F) = 6 THEN
               #inState := #inState + 1;
           ELSE
               #q_xError := TRUE;
               #inErrorState := #inState;
               #inState := 100;
           END_IF;
           // ******************************************************************************************************

